FUNCTION "LGF_IntToString" : String   // FC10046, SCL
{ S7_Optimized_Access := 'TRUE' }
VERSION : 0.1
   VAR_INPUT
      intValue : DInt;   // Integer value to convert
   END_VAR
   VAR_TEMP
      tempString : String;   // Temp string
   END_VAR
   // Ret_Val : Converted integer
BEGIN
   //=============================================================================
   // Siemens AG
   // (c)Copyright 2017
   //-----------------------------------------------------------------------------
   // Library:       LGF (Library General Functions)
   // Tested with:   CPU1212C DC/DC/DC FW:V4.2
   // Engineering:   TIA Portal V14 SP1 Upd 5
   // Restrictions:  -
   // Requirements:  PLC (S7-1200 / S7-1500)
   // Functionality: This function converts a integer value to a string
   //-----------------------------------------------------------------------------
   // Change log table:
   // Version  Date        In charge / Changes applied
   // 01.00.00 04.07.2018  Siemens Industry Online Support
   //                      First released version
   // 01.00.01 17.08.2018  Siemens Industry Online Support
   //                      Upgrade: TIA V15 Update 2
   // 01.00.02 23.11.2018  Siemens Industry Online Support
   //                      Upgrade: TIA V15.1
   //=============================================================================

   // Convert integer to string
   #tempString := DINT_TO_STRING(#intValue);

   // Delete padding before number
   WHILE (FIND(IN1 := #tempString, IN2 := ' ') <> 0) DO
     #tempString := DELETE(IN := #tempString, L := 1, P := 1);
   END_WHILE;

   // Output string
   #LGF_IntToString := #tempString;
END_FUNCTION

FUNCTION "LGF_UnixTimeToDTL" : DTL   // FC10047, SCL
{ S7_Optimized_Access := 'TRUE' }
VERSION : 0.1
   VAR_INPUT
      timeUnix : DInt;   // Unix time to convert
   END_VAR
   VAR_OUTPUT
      error : Bool;   // Error = TRUE: Time is outside of allowed range
   END_VAR
   VAR_TEMP
      tempDate : DInt;   // Temporary Date value
      tempTime : DInt;   // Temporary Time value
      tempDTL : DTL;   // Temporary DTL value
   END_VAR
   // Ret_Val : Converted time in DTL
   VAR CONSTANT
      DELTA_1970_1990 : DInt := 631_152_000;   // Delta between 1970-1-1 and 1990-1-1 in seconds (IEC Time Base)
      SEC_PER_DAY : DInt := 86400;   // 86400 seconds in 1 day
   END_VAR
BEGIN
   //=============================================================================
   // Siemens AG
   // (c)Copyright 2017
   //-----------------------------------------------------------------------------
   // Library:       LGF (Library General Functions)
   // Tested with:   CPU1212C DC/DC/DC FW:V4.2
   // Engineering:   TIA Portal V15
   // Restrictions:  -
   // Requirements:  PLC (S7-1200 / S7-1500)
   // Functionality: This function converts Unix time to DTL
   //-----------------------------------------------------------------------------
   // Change log table:
   // Version  Date        In charge / Changes applied
   // 01.00.00 16.10.2018  Siemens Industry Online Support
   //                      First released version
   //=============================================================================

   #error := FALSE;

   // Check if timeUnix less than 01.01.1990
   IF (#timeUnix < #DELTA_1970_1990)
   THEN
     #error := TRUE;
     #LGF_UnixTimeToDTL := DTL#1990-01-01-00:00:00;
     RETURN;
   END_IF;

   // Convert date
   #tempDate := (#timeUnix - #DELTA_1970_1990) / #SEC_PER_DAY;
   #tempDTL := DATE_TO_DTL(DINT_TO_DATE(#tempDate));

   // Convert time
   #tempTime := #timeUnix - #DELTA_1970_1990 - (#tempDate * #SEC_PER_DAY);
   #tempDTL.HOUR := DINT_TO_USINT(#tempTime / 3600);
   #tempDTL.MINUTE := DINT_TO_USINT(#tempTime MOD 3600 / 60);
   #tempDTL.SECOND := DINT_TO_USINT(#tempTime MOD 60);

   // Output date and time
   #LGF_UnixTimeToDTL := #tempDTL;
END_FUNCTION

FUNCTION "LGF_DTLToUnixTime" : DInt   // FC10048, SCL
{ S7_Optimized_Access := 'TRUE' }
VERSION : 0.1
   VAR_INPUT
      timeDTL : DTL;   // Time in DTL to convert
   END_VAR
   VAR_OUTPUT
      error : Bool;   // Error = TRUE: Time is outside of allowed range
   END_VAR
   // Ret_Val : Converted Unix time
   VAR CONSTANT
      DELTA_1970_1990 : DInt := 631_152_000;   // Delta between 1970-1-1 and 1990-1-1 in seconds (IEC Time Base)
      SEC_PER_DAY : DInt := 86400;   // 86400 seconds in 1 day
   END_VAR
BEGIN
   //=============================================================================
   // Siemens AG
   // (c)Copyright 2017
   //-----------------------------------------------------------------------------
   // Library:       LGF (Library General Functions)
   // Tested with:   CPU1212C DC/DC/DC FW:V4.2
   // Engineering:   TIA Portal V15
   // Restrictions:  -
   // Requirements:  PLC (S7-1200 / S7-1500)
   // Functionality: This function converts DTL to Unix time
   //-----------------------------------------------------------------------------
   // Change log table:
   // Version  Date        In charge / Changes applied
   // 01.00.00 16.10.2018  Siemens Industry Online Support
   //                      First released version
   //=============================================================================

   #error := FALSE;

   // Check if timeUnix less than 01.01.1990
   IF (#timeDTL < DTL#1990-01-01-00:00:00)
   THEN
     #error := TRUE;
     #LGF_DTLToUnixTime := 0;
     RETURN;
   END_IF;

   // Convert System Time (UTC) to UNIX time
   #LGF_DTLToUnixTime := (DATE_TO_DINT(DTL_TO_DATE(#timeDTL)) * #SEC_PER_DAY)
                       + (TOD_TO_DINT(DTL_TO_TOD(#timeDTL)) / 1000)
                       + #DELTA_1970_1990;
END_FUNCTION

// folder: Phisical_functions/LGF/7 Signal generators

FUNCTION_BLOCK "LGF_Frequency"   // FB10024, SCL
{ S7_Optimized_Access := 'TRUE' }
   VAR_INPUT
      frequency : Real;   // Input in Hz
      pulsePauseRatio : Real := 1.0;   // Pulse pause ratio
   END_VAR
   VAR_OUTPUT
      clock : Bool;   // -
      countdown : Time;   // -
   END_VAR
   VAR
      instTofTimePulse : TOF_TIME;   // -
      instTofTimePause : TOF_TIME;   // -
      statFrequency : Real;   // -
      statTimePeriod : Time;   // -
      statTimePulse : Time;   // -
      statTimePause : Time;   // -
      statPulsePauseRatio : Real;   // -
   END_VAR
   VAR_TEMP
      tempPulseRate : Real;   // -
      tempPauseRate : Real;   // -
   END_VAR
   VAR CONSTANT
      NULL : Real := 0.0;   // -
   END_VAR
BEGIN
   //=============================================================================
   // SIEMENS AG
   // (c)Copyright 2017
   //-----------------------------------------------------------------------------
   // Library:       LGF (Library General Functions)
   // Tested with:   CPU1214C DC/DC/DC FW:V4.2
   // Engineering:   TIA Portal V14
   // Restrictions:  -
   // Requirements:  PLC (S7-1200, S7-1500)
   // Functionality: Generates frequency signal
   //-----------------------------------------------------------------------------
   // Change log table:
   // Version  Date        Expert in charge / Changes applied
   // 01.00.00 19.08.2015  Siemens Industry Online Support
   //                      First released version
   // 01.01.00 25.05.2016  Siemens Industry Online Support
   //                      New function: pulse pause ratio
   // 01.01.01 26.05.2016  Siemens Industry Online Support
   //                      Add comments
   // 01.01.02 02.01.2017  Siemens Industry Online Support
   //                      Upgrade: TIA Portal V14 Update 1
   // 01.01.03 17.08.2018  Siemens Industry Online Support
   //                      Upgrade: TIA V15 Update 2
   // 01.01.04 23.11.2018  Siemens Industry Online Support
   //                      Upgrade: TIA V15.1
   //=============================================================================

   IF (#frequency <= #NULL) OR (#pulsePauseRatio <= #NULL)  // If input is <= 0.0 : block is off
   THEN
     #clock := FALSE;
     #countdown := t#0s;
   ELSE
     // assign frequency and pulse pause ratio one time 
     IF #statFrequency <> #frequency OR #statPulsePauseRatio <> #pulsePauseRatio THEN
       RESET_TIMER(TIMER := #instTofTimePause);
       RESET_TIMER(TIMER := #instTofTimePulse);

       #tempPulseRate := #pulsePauseRatio / (#pulsePauseRatio + 1); // Calculate pulse rate   
       #tempPauseRate := 1.0 - #tempPulseRate;                      // Calculate pause rate   
       #statTimePeriod := UDINT_TO_TIME(REAL_TO_UDINT((1000.0 / #frequency)));                 // Calculate period time 
       #statTimePulse := UDINT_TO_TIME(REAL_TO_UDINT((1000.0 * #tempPulseRate / #frequency))); // Calculate pulse time   
       #statTimePause := UDINT_TO_TIME(REAL_TO_UDINT((1000.0 * #tempPauseRate / #frequency))); // Calculate pause time
       #statFrequency := #frequency;
       #statPulsePauseRatio := #pulsePauseRatio;
     END_IF;

     // TOF_off expired >> Start again
     #instTofTimePulse(IN := NOT #instTofTimePause.Q,
                       PT := #statTimePulse);
     #countdown := #statTimePulse - #instTofTimePulse.ET;

     #instTofTimePause(IN := #instTofTimePulse.Q,
                       PT := #statTimePause);

     IF #countdown = t#0s THEN
       #countdown := #statTimePause - #instTofTimePause.ET;
     END_IF;

     #clock := #instTofTimePulse.Q; // Assign ouptut 
   END_IF;
END_FUNCTION_BLOCK

FUNCTION_BLOCK "LGF_Impulse"   // FB10025, SCL
{ S7_Optimized_Access := 'TRUE' }
   VAR_INPUT
      frequency : Real;   // Frequnency in Hz
   END_VAR
   VAR_OUTPUT
      impulse : Bool;   // Impulse output
      countdown : Time;   // -
   END_VAR
   VAR
      instTofTimePulse : TOF_TIME;
      statFrequency : Real;
      statTimePulse : Time;
   END_VAR
   VAR_TEMP
      tempImpulse : Bool;
      tempCountdown : Time;
   END_VAR
BEGIN
   //=============================================================================
   // SIEMENS AG
   // (c)Copyright 2017
   //-----------------------------------------------------------------------------
   // Library:       LGF (Library General Functions)
   // Tested with:   CPU1212C DC/DC/DC FW:V4.1
   // Engineering:   TIA Portal V14 Update 1
   // Restrictions:  -
   // Requirements:  PLC (S7-1200 / S7-1500)
   // Functionality: This fuction block generates impulses in the given frequency 
   //-----------------------------------------------------------------------------
   // Change log table:
   // Version  Date        Expert in charge / Changes applied
   // 01.00.00 19.08.2015  Siemens Industry Online Support
   //                      First released version
   // 01.01.01 16.06.2015  Siemens Industry Online Support
   //                      LGF_Impulse calls new LGF_Frequency V1.1.1
   // 01.01.02 02.01.2017  Siemens Industry Online Support
   //                      Upgrade: TIA Portal V14 Update 1
   // 01.02.00 02.02.2017  Siemens Industry Online Support
   //                      Code optimization: no call of LGF_Frequency
   //                      Fix at output "countdown"
   // 01.02.01 17.08.2018  Siemens Industry Online Support
   //                      Upgrade: TIA V15 Update 2
   // 01.02.02 23.11.2018  Siemens Industry Online Support
   //                      Upgrade: TIA V15.1
   //=============================================================================

   IF #frequency <= 0.0 THEN
     #tempImpulse := FALSE;
     #tempCountdown := t#0s;

   ELSE
     // Assign frequency
     #statTimePulse := t#1000s / TRUNC(#frequency * 1000);
     #statFrequency := #frequency;

     // Assign impulse
     #tempImpulse := NOT #instTofTimePulse.Q;

     // Time pulse expired >> Start again
     #instTofTimePulse(IN := NOT #instTofTimePulse.Q,
                       PT := #statTimePulse);

     // Assign countdown
     #tempCountdown := #statTimePulse - #instTofTimePulse.ET;
   END_IF;

   // Write outputs
   #impulse := #tempImpulse;
   #countdown := #tempCountdown;
END_FUNCTION_BLOCK

FUNCTION_BLOCK "LGF_SawTooth"   // FB10026, SCL
{ S7_Optimized_Access := 'TRUE' }
   VAR_INPUT
      startValue : Int;
      timeRange : Time;
      incrementRange : Int;
      numberSteps : Int;
      endlessSteps : Bool;
      restart : Bool;
   END_VAR
   VAR_OUTPUT
      value : Int;
   END_VAR
   VAR
      statStartValue : Int;   // start value of the saw tooth
      statTimeRange : Time;   // time of one period
      statIncrementRange : Int;   // difference from one to another value
      statNumberSteps : Int;   // number of steps
      statEndlessSteps : Bool;
      statCurrentStep : Int;
      statPrevValue : Int;
      statFirstRun : Bool := TRUE;
      statEndlessOn : Bool;
      statStartTimer : Bool;
      statTimerFinished : Bool;
      instTimer : TON_TIME;
      statActValue : Int;
   END_VAR
BEGIN
   //=============================================================================
   // SIEMENS AG
   // (c)Copyright 2017
   //-----------------------------------------------------------------------------
   // Library:       LGF(Library General Functions)
   // Tested with:   CPU1212C DC/DC/DC FW:V4.2
   // Engineering:   TIA Portal V14 Update 1
   // Restrictions:  -
   // Requirements:  PLC (S7-1200 / S7-1500)
   // Functionality: Saw tooth generator
   //-----------------------------------------------------------------------------
   // Change log table:
   // Version  Date        Expert in charge / Changes applied
   // 01.00.00 19.08.2015  Siemens Industry Online Support
   //                      First released version
   // 01.00.01 02.11.2015  Siemens Industry Online Support
   //                      Bug fix
   // 01.00.02 02.01.2017  Siemens Industry Online Support
   //                      Upgrade: TIA Portal V14 Update 1
   // 01.00.03 17.08.2018  Siemens Industry Online Support
   //                      Upgrade: TIA V15 Update 2
   // 01.00.04 23.11.2018  Siemens Industry Online Support
   //                      Upgrade: TIA V15.1
   //=============================================================================

   // Initialization for the first call or reset complete function
   IF (#statFirstRun = TRUE)
     OR (#restart = TRUE) THEN

     // Copy all input parameter to static values
     #statStartValue := #startValue;
     #statTimeRange := #timeRange;
     #statIncrementRange := #incrementRange;
     #statNumberSteps := #numberSteps;
     #statEndlessSteps := #endlessSteps;

     // Reset static values
     #statActValue := #statStartValue;
     #statStartTimer := TRUE;
     #statCurrentStep := 0;
     #statFirstRun := FALSE;
   END_IF;

   // Calculation of a new values if the time base is up
   IF #statTimerFinished = TRUE
     AND (#restart = FALSE) THEN

     #statActValue := #statActValue + #statIncrementRange;
     #statCurrentStep := #statCurrentStep + 1;

     // If a defined number of steps must be performed 
     IF (#statEndlessSteps = FALSE) THEN

       // Restart with start value if number of steps is reached
       IF #statCurrentStep > #statNumberSteps THEN

         #statCurrentStep := 0;
         #statActValue := #statStartValue;
       END_IF;

       // If endless is on the step counter is resetted  
     ELSE

       #statEndlessOn := TRUE;
       #statCurrentStep := 0;
     END_IF;

     #statStartTimer := FALSE; // Reset the time base
   END_IF;

   // Call a times as basis of the step range
   #instTimer(IN := #statStartTimer,
              PT := #statTimeRange,
              Q => #statTimerFinished);

   // Start the timer
   #statStartTimer := TRUE;

   // Write Output, if restart is active output value = 0
   IF (#restart = TRUE) THEN
     #statActValue := #startValue;
   END_IF;

   #value := #statActValue;
END_FUNCTION_BLOCK

FUNCTION_BLOCK "LGF_SinusCI"   // FB10027, SCL
{ S7_Optimized_Access := 'TRUE' }
VERSION : 0.1
   VAR_INPUT
      amplitude : Real := 0.0;   // Amplitude
      offset : Real := 1000.0;   // Offset
      periodeMS : UDInt := 1000;   // Periode in milliseconds
      callOB : OB_Cyclic;   // Call OB
      reset : Bool;   // Reset values
   END_VAR
   VAR_OUTPUT
      sinusValues : Real;   // Calculated Sinus values
      error : Bool;   // "0" = no error; "1" = error
      statusID : UInt;   // Error source
      status : Word;   // Status and error codes
   END_VAR
   VAR
      statRad : Real;   // Size of an angle in radians
      statCounter : UDInt;   // Counter value
   END_VAR
   VAR_TEMP
      tempCycleTime : UDInt;   // Temp cycle time from CallOB
      tempCyclePhase : UDInt;   // Temp cycle phase from CallOB
      tempCycleStatus : Word;   // Temp cycle status from CallOB
      tempReadTimeStatus : Int;   // Return value of QRY_CINT
   END_VAR
   VAR CONSTANT
      PI : Real := 3.141593;   // PI
      NO_ERROR : Word := 16#0000;   // Status no error
      OB_UNAVAILABLE : Word := 16#8200;   // Status OB not available
      ERROR_IN_THIS_BLOCK : UInt := 1;   // Error ID local error
      ERROR_QRY_CINT : UInt := 2;   // Error ID error in function QRY_CINT
   END_VAR
BEGIN
   //=============================================================================
   // Siemens AG
   // (c)Copyright 2017
   //-----------------------------------------------------------------------------
   // Library:       LGF (Library General Functions)
   // Tested with:   CPU1212C DC/DC/DC FW:V4.2
   // Engineering:   TIA Portal V15 Upd 2
   // Restrictions:  -
   // Requirements:  PLC (S7-1200 / S7-1500)
   // Functionality: This function generates a sinus signal
   //-----------------------------------------------------------------------------
   // Change log table:
   // Version  Date        In charge/Changes applied
   // 01.00.00 03.07.2018  Siemens Industry Online Support
   //                      First released version
   // 01.00.01 17.08.2018  Siemens Industry Online Support
   //                      Upgrade: TIA V15 Update 2
   // 01.00.02 23.11.2018  Siemens Industry Online Support
   //                      Upgrade: TIA V15.1
   //-----------------------------------------------------------------------------
   //Status Codes: -
   //=============================================================================

   // Initialize
   #error := FALSE;
   #statusID := #ERROR_IN_THIS_BLOCK;
   #status := #NO_ERROR;

   // get sample time, according to the cyclic interrupt OB number
   #tempReadTimeStatus := QRY_CINT(OB_NR := #callOB, CYCLE => #tempCycleTime,
                                   PHASE => #tempCyclePhase, STATUS => #tempCycleStatus);

   // Generate error message of the QRY_CINT function
   IF (#tempReadTimeStatus <> 0)
   THEN
     #error := TRUE;
     #statusID := #ERROR_QRY_CINT;
     #status := INT_TO_WORD(#tempReadTimeStatus);
     RETURN;
   END_IF;

   // Generate error message when OB unavailable
   IF (#tempCycleStatus = 16#0000)
   THEN
     #error := TRUE;
     #statusID := #ERROR_IN_THIS_BLOCK;
     #status := #OB_UNAVAILABLE;
     RETURN;
   END_IF;

   IF (#reset = TRUE)
   THEN
     #statCounter := 0;
     #sinusValues := 0;
   ELSE
     // Increment Counter with each call of "OB_Cyclic_interrupt"
     #statCounter := #statCounter + (#tempCycleTime) / 1000;
     #statCounter := #statCounter MOD (#periodeMS);

     #statRad := UDINT_TO_REAL(#statCounter) * 2.0 * #PI / (UDINT_TO_REAL(#periodeMS));

     #sinusValues := SIN(#statRad) * #amplitude + #offset;
   END_IF;
END_FUNCTION_BLOCK

FUNCTION_BLOCK "LGF_CosinusCI"   // FB10028, SCL
{ S7_Optimized_Access := 'TRUE' }
VERSION : 0.1
   VAR_INPUT
      amplitude : Real := 0.0;   // Amplitude
      offset : Real := 1000.0;   // Offset
      periodeMS : UDInt := 1000;   // Periode in milliseconds
      callOB : OB_Cyclic;   // Call OB
      reset : Bool;   // Reset values
   END_VAR
   VAR_OUTPUT
      cosinusValues : Real;   // Calculated Cosinus values
      error : Bool;   // "0" = no error; "1" = error
      statusID : UInt;   // Error source
      status : Word;   // Status and error codes
   END_VAR
   VAR
      statRad : Real;   // Size of an angle in radians
      statCounter : UDInt;   // Counter value
   END_VAR
   VAR_TEMP
      tempCycleTime : UDInt;   // Temp cycle time from CallOB
      tempCyclePhase : UDInt;   // Temp cycle phase from CallOB
      tempCycleStatus : Word;   // Temp cycle status from CallOB
      tempReadTimeStatus : Int;   // Return value of QRY_CINT
   END_VAR
   VAR CONSTANT
      PI : Real := 3.141593;   // PI
      NO_ERROR : Word := 16#0000;   // Status no error
      OB_UNAVAILABLE : Word := 16#8200;   // Status OB not available
      ERROR_IN_THIS_BLOCK : UInt := 1;   // Error ID local error
      ERROR_QRY_CINT : UInt := 2;   // Error ID error in function QRY_CINT
   END_VAR
BEGIN
   //=============================================================================
   // Siemens AG
   // (c)Copyright 2017
   //-----------------------------------------------------------------------------
   // Library:       LGF (Library General Functions)
   // Tested with:   CPU1212C DC/DC/DC FW:V4.2
   // Engineering:   TIA Portal V15 Upd 2
   // Restrictions:  -
   // Requirements:  PLC (S7-1200 / S7-1500)
   // Functionality: This function generates a cosinus signal
   //-----------------------------------------------------------------------------
   // Change log table:
   // Version  Date        In charge/Changes applied
   // 01.00.00 03.07.2018  Siemens Industry Online Support
   //                      First released version
   // 01.00.01 17.08.2018  Siemens Industry Online Support
   //                      Upgrade: TIA V15 Update 2
   // 01.00.02 23.11.2018  Siemens Industry Online Support
   //                      Upgrade: TIA V15.1
   //-----------------------------------------------------------------------------
   //Status Codes: -
   //=============================================================================

   // Initialize
   #error := FALSE;
   #statusID := #ERROR_IN_THIS_BLOCK;
   #status := #NO_ERROR;

   // get sample time, according to the cyclic interrupt OB number
   #tempReadTimeStatus := QRY_CINT(OB_NR := #callOB, CYCLE => #tempCycleTime,
                                   PHASE => #tempCyclePhase, STATUS => #tempCycleStatus);

   // Generate error message of the QRY_CINT function
   IF (#tempReadTimeStatus <> 0)
   THEN
     #error := TRUE;
     #statusID := #ERROR_QRY_CINT;
     #status := INT_TO_WORD(#tempReadTimeStatus);
     RETURN;
   END_IF;

   // Generate error message when OB unavailable
   IF (#tempCycleStatus = 16#0000)
   THEN
     #error := TRUE;
     #statusID := #ERROR_IN_THIS_BLOCK;
     #status := #OB_UNAVAILABLE;
     RETURN;
   END_IF;

   IF (#reset = TRUE) 
   THEN
     #statCounter := 0;
     #cosinusValues := 0;
   ELSE
     // Increment Counter with each call of "OB_Cyclic_interrupt"
     #statCounter := #statCounter + (#tempCycleTime) / 1000;
     #statCounter := #statCounter MOD (#periodeMS);

     #statRad := UDINT_TO_REAL(#statCounter) * 2.0 * #PI / (UDINT_TO_REAL(#periodeMS));

     #cosinusValues := COS(#statRad) * #amplitude + #offset;
   END_IF;
END_FUNCTION_BLOCK

FUNCTION_BLOCK "LGF_RectangleCI"   // FB10029, SCL
{ S7_Optimized_Access := 'TRUE' }
VERSION : 0.1
   VAR_INPUT
      amplitude : Real := 0.0;   // Amplitude
      offset : Real := 1000.0;   // Offset
      periodeMS : UDInt := 1000;   // Periode in milliseconds
      callOB : OB_Cyclic;   // Call OB
      reset : Bool;   // Reset values
   END_VAR
   VAR_OUTPUT
      rectangleValues : Real;   // Calculated rectangle values
      error : Bool;   // "0" = no error; "1" = error
      statusID : UInt;   // Error source
      status : Word;   // Status and error codes
   END_VAR
   VAR
      statRad : Real;   // Size of an angle in radians
      statCounter : UDInt;   // Counter value
   END_VAR
   VAR_TEMP
      tempCycleTime : UDInt;   // Temp cycle time from CallOB
      tempCyclePhase : UDInt;   // Temp cycle phase from CallOB
      tempCycleStatus : Word;   // Temp cycle status from CallOB
      tempReadTimeStatus : Int;   // Return value of QRY_CINT
   END_VAR
   VAR CONSTANT
      PI : Real := 3.141593;   // PI
      NO_ERROR : Word := 16#0000;   // Status no error
      OB_UNAVAILABLE : Word := 16#8200;   // Status OB not available
      ERROR_IN_THIS_BLOCK : UInt := 1;   // Error ID local error
      ERROR_QRY_CINT : UInt := 2;   // Error ID error in function QRY_CINT
   END_VAR
BEGIN
   //=============================================================================
   // Siemens AG
   // (c)Copyright 2017
   //-----------------------------------------------------------------------------
   // Library:       LGF (Library General Functions)
   // Tested with:   CPU1212C DC/DC/DC FW:V4.2
   // Engineering:   TIA Portal V15 Upd 2
   // Restrictions:  -
   // Requirements:  PLC (S7-1200 / S7-1500)
   // Functionality: This function generates a rectangle signal
   //-----------------------------------------------------------------------------
   // Change log table:
   // Version  Date        In charge/Changes applied
   // 01.00.00 03.07.2018  Siemens Industry Online Support
   //                      First released version
   // 01.00.01 17.08.2018  Siemens Industry Online Support
   //                      Upgrade: TIA V15 Update 2
   // 01.00.02 23.11.2018  Siemens Industry Online Support
   //                      Upgrade: TIA V15.1
   //-----------------------------------------------------------------------------
   //Status Codes: -
   //=============================================================================

   // Initialize
   #error := FALSE;
   #statusID := #ERROR_IN_THIS_BLOCK;
   #status := #NO_ERROR;

   // get sample time, according to the cyclic interrupt OB number
   #tempReadTimeStatus := QRY_CINT(OB_NR := #callOB, CYCLE => #tempCycleTime,
                                   PHASE => #tempCyclePhase, STATUS => #tempCycleStatus);

   // Generate error message of the QRY_CINT function
   IF (#tempReadTimeStatus <> 0)
   THEN
     #error := TRUE;
     #statusID := #ERROR_QRY_CINT;
     #status := INT_TO_WORD(#tempReadTimeStatus);
     RETURN;
   END_IF;

   // Generate error message when OB unavailable
   IF (#tempCycleStatus = 16#0000)
   THEN
     #error := TRUE;
     #statusID := #ERROR_IN_THIS_BLOCK;
     #status := #OB_UNAVAILABLE;
     RETURN;
   END_IF;

   IF (#reset = TRUE) 
   THEN
     #statCounter := 0;
     #rectangleValues := 0;
   ELSE
     // Increment Counter with each call of "OB_Cyclic_interrupt"
     #statCounter := #statCounter + (#tempCycleTime) / 1000;
     #statCounter := #statCounter MOD (#periodeMS);

     IF (#statCounter <= (#periodeMS / 2))
     THEN
       #rectangleValues := #offset + #amplitude;
     ELSE
       #rectangleValues := #offset - #amplitude;
     END_IF;
   END_IF;
END_FUNCTION_BLOCK

FUNCTION_BLOCK "LGF_TriangleCI"   // FB10030, SCL
{ S7_Optimized_Access := 'TRUE' }
VERSION : 0.1
   VAR_INPUT
      amplitude : Real := 0.0;   // Amplitude
      offset : Real := 1000.0;   // Offset
      periodeMS : UDInt := 1000;   // Periode in milliseconds
      callOB : OB_Cyclic;   // Call OB
      reset : Bool;   // Reset values
   END_VAR
   VAR_OUTPUT
      triangleValues : Real;   // Calculated triangle values
      error : Bool;   // "0" = no error; "1" = error
      statusID : UInt;   // Error source
      status : Word;   // Status and error codes
   END_VAR
   VAR
      statRad : Real;   // Size of an angle in radians
      statCounter : UDInt;   // Counter value
   END_VAR
   VAR_TEMP
      tempCycleTime : UDInt;   // Temp cycle time from CallOB
      tempCyclePhase : UDInt;   // Temp cycle phase from CallOB
      tempCycleStatus : Word;   // Temp cycle status from CallOB
      tempReadTimeStatus : Int;   // Return value of QRY_CINT
   END_VAR
   VAR CONSTANT
      PI : Real := 3.141593;   // PI
      NO_ERROR : Word := 16#0000;   // Status no error
      OB_UNAVAILABLE : Word := 16#8200;   // Status OB not available
      ERROR_IN_THIS_BLOCK : UInt := 1;   // Error ID local error
      ERROR_QRY_CINT : UInt := 2;   // Error ID error in function QRY_CINT
   END_VAR
BEGIN
   //=============================================================================
   // Siemens AG
   // (c)Copyright 2017
   //-----------------------------------------------------------------------------
   // Library:       LGF (Library General Functions)
   // Tested with:   CPU1212C DC/DC/DC FW:V4.2
   // Engineering:   TIA Portal V15 Upd 2
   // Restrictions:  -
   // Requirements:  PLC (S7-1200 / S7-1500)
   // Functionality: This function generates a rectangle signal
   //-----------------------------------------------------------------------------
   // Change log table:
   // Version  Date        In charge/Changes applied
   // 01.00.00 03.07.2018  Siemens Industry Online Support
   //                      First released version
   // 01.00.01 17.08.2018  Siemens Industry Online Support
   //                      Upgrade: TIA V15 Update 2
   // 01.00.02 23.11.2018  Siemens Industry Online Support
   //                      Upgrade: TIA V15.1
   //-----------------------------------------------------------------------------
   //Status Codes: -
   //=============================================================================

   // Initialize
   #error := FALSE;
   #statusID := #ERROR_IN_THIS_BLOCK;
   #status := #NO_ERROR;

   // get sample time, according to the cyclic interrupt OB number
   #tempReadTimeStatus := QRY_CINT(OB_NR := #callOB, CYCLE => #tempCycleTime,
                                   PHASE => #tempCyclePhase, STATUS => #tempCycleStatus);

   // Generate error message of the QRY_CINT function
   IF (#tempReadTimeStatus <> 0)
   THEN
     #error := TRUE;
     #statusID := #ERROR_QRY_CINT;
     #status := INT_TO_WORD(#tempReadTimeStatus);
     RETURN;
   END_IF;

   // Generate error message when OB unavailable
   IF #tempCycleStatus = 16#0000 THEN
     #error := TRUE;
     #statusID := #ERROR_IN_THIS_BLOCK;
     #status := #OB_UNAVAILABLE;
     RETURN;
   END_IF;

   IF (#reset = TRUE) 
   THEN
     #statCounter := 0;
     #triangleValues := 0;
   ELSE
     // Increment Counter with each call of "OB_Cyclic_interrupt"
     #statCounter := #statCounter + (#tempCycleTime) / 1000;
     #statCounter := #statCounter MOD (#periodeMS);

     IF (#statCounter <= (#periodeMS / 2))
     THEN
       #triangleValues := 4.0 * #amplitude /  UDINT_TO_REAL(#periodeMS) * UDINT_TO_REAL(#statCounter)  - #amplitude + #offset;
     ELSE
       #triangleValues := -4.0 * #amplitude / UDINT_TO_REAL(#periodeMS) * UDINT_TO_REAL(#statCounter) + 3 * #amplitude + #offset;
     END_IF;
   END_IF;
END_FUNCTION_BLOCK

FUNCTION_BLOCK "LGF_SawToothCI"   // FB10031, SCL
{ S7_Optimized_Access := 'TRUE' }
VERSION : 0.1
   VAR_INPUT
      amplitude : Real := 0.0;   // Amplitude
      offset : Real := 1000.0;   // Offset
      periodeMS : UDInt := 1000;   // Periode in milliseconds
      callOB : OB_Cyclic;   // Call OB
      reset : Bool;   // Reset values
   END_VAR
   VAR_OUTPUT
      sawToothValues : Real;   // Calculated saw tooth values
      error : Bool;   // "0" = no error; "1" = error
      statusID : UInt;   // Error source
      status : Word;   // Status and error codes
   END_VAR
   VAR
      statRad : Real;   // Size of an angle in radians
      statCounter : UDInt;   // Counter value
   END_VAR
   VAR_TEMP
      tempCycleTime : UDInt;   // Temp cycle time from CallOB
      tempCyclePhase : UDInt;   // Temp cycle phase from CallOB
      tempCycleStatus : Word;   // Temp cycle status from CallOB
      tempReadTimeStatus : Int;   // Return value of QRY_CINT
   END_VAR
   VAR CONSTANT
      PI : Real := 3.141593;   // PI
      NO_ERROR : Word := 16#0000;   // Status no error
      OB_UNAVAILABLE : Word := 16#8200;   // Status OB not available
      ERROR_IN_THIS_BLOCK : UInt := 1;   // Error ID local error
      ERROR_QRY_CINT : UInt := 2;   // Error ID error in function QRY_CINT
   END_VAR
BEGIN
   //=============================================================================
   // Siemens AG
   // (c)Copyright 2017
   //-----------------------------------------------------------------------------
   // Library:       LGF (Library General Functions)
   // Tested with:   CPU1212C DC/DC/DC FW:V4.2
   // Engineering:   TIA Portal V15 Upd 2
   // Restrictions:  -
   // Requirements:  PLC (S7-1200 / S7-1500)
   // Functionality: This function generates a rectangle signal
   //-----------------------------------------------------------------------------
   // Change log table:
   // Version  Date        In charge/Changes applied
   // 01.00.00 03.07.2018  Siemens Industry Online Support
   //                      First released version
   // 01.00.01 17.08.2018  Siemens Industry Online Support
   //                      Upgrade: TIA V15 Update 2
   // 01.00.02 23.11.2018  Siemens Industry Online Support
   //                      Upgrade: TIA V15.1
   //-----------------------------------------------------------------------------
   //Status Codes: -
   //=============================================================================

   // Initialize
   #error := FALSE;
   #statusID := #ERROR_IN_THIS_BLOCK;
   #status := #NO_ERROR;

   // get sample time, according to the cyclic interrupt OB number
   #tempReadTimeStatus := QRY_CINT(OB_NR := #callOB, CYCLE => #tempCycleTime,
                                   PHASE => #tempCyclePhase, STATUS => #tempCycleStatus);

   // Generate error message of the QRY_CINT function
   IF (#tempReadTimeStatus <> 0)
   THEN
     #error := TRUE;
     #statusID := #ERROR_QRY_CINT;
     #status := INT_TO_WORD(#tempReadTimeStatus);
     RETURN;
   END_IF;

   // Generate error message when OB unavailable
   IF (#tempCycleStatus = 16#0000)
   THEN
     #error := TRUE;
     #statusID := #ERROR_IN_THIS_BLOCK;
     #status := #OB_UNAVAILABLE;
     RETURN;
   END_IF;

   IF (#reset = TRUE)
   THEN
     #statCounter := 0;
     #sawToothValues := 0;
   ELSE
     // Increment Counter with each call of "OB_Cyclic_interrupt"
     #statCounter := #statCounter + (#tempCycleTime) / 1000;
     #statCounter := #statCounter MOD (#periodeMS);

     #sawToothValues := 2.0 * #amplitude / UDINT_TO_REAL(#periodeMS) * UDINT_TO_REAL(#statCounter) - #amplitude + #offset;

   END_IF;
END_FUNCTION_BLOCK

// folder: Phisical_functions/LGF/8 Technology operations

FUNCTION_BLOCK "LGF_LimRateOfChangeBasic"   // FB10032, SCL
{ S7_Optimized_Access := 'TRUE' }
VERSION : 0.1
   VAR_INPUT
      inputValue : Real;   // Input Value/ setpoint
      setRateLim : Real;   // rate of change limitation (1/second)
      defaultOutValue : Real;   // default output value
      onDefaultOutValue : Bool;   // default output value on (outputValue=defaultOutValue)
      callOB : OB_Cyclic;   // cyclic interrupt OB
   END_VAR
   VAR_OUTPUT
      outputValue : Real;   // output value
      error : Bool;   // "0" = no error; "1" = error
      statusID : UInt;   // Error destination: "1" = LGFLimRateOfChangeBasic; "2" = QRY_CINT
      status : Word;   // status and error codes
   END_VAR
   VAR
      statPrevTime : DTL;   // -
      statPrevOut : Real;   // -
   END_VAR
   VAR_TEMP
      tempCycleTime : UDInt;   // -
      tempCylcePhase : UDInt;   // -
      tempCycleStatus : Word;   // -
      tempDeltaTime : Time;   // -
      tempCycleTimeReal : Real;   // -
      tempReadTimeStatus : Int;   // -
      tempOut : Real;   // -
   END_VAR
   VAR CONSTANT
      NO_ERROR : Word := 16#0000;   // -
      INIT_VALUE : Word := 16#7000;   // -
      OB_UNAVAILABLE : Word := 16#8200;   // -
      NEG_RATE_LIM : Word := 16#8201;   // -
      ERROR_IN_THIS_BLOCK : UInt := 1;   // -
      ERROR_QRY_CINT : UInt := 2;   // -
   END_VAR
BEGIN
   //=============================================================================
   // Siemens AG
   // (c)Copyright 2017
   //-----------------------------------------------------------------------------
   // Library:       LGF(Library General Functions)
   // Tested with:   CPU1212C DC/DC/DC FW:V4.2
   // Engineering:   TIA Portal V14 Update 1
   // Restrictions:  only callable in a cyclic interrupt OB
   // Requirements:  PLC (S7-1200 / S7-1500)
   // Functionality: This function block generates a ramp function from a step function.
   //-----------------------------------------------------------------------------
   // Change log table:
   // Version  Date        In charge / Changes applied
   // 01.00.00 21.06.2016  Siemens Industry Online Support
   //                      First released version
   // 01.00.01 02.01.2017  Siemens Industry Online Support
   //                      Upgrade: TIA Portal V14 Update 1
   // 01.00.02 17.08.2018  Siemens Industry Online Support
   //                      Upgrade: TIA V15 Update 2
   // 01.00.03 23.11.2018  Siemens Industry Online Support
   //                      Upgrade: TIA V15.1
   //-----------------------------------------------------------------------------
   //Status Codes:
   // 16#0000:  No errors
   // 16#7000:  Initial value
   // 16#8200:  Call OB unavailable
   // 16#8201:  Negativ value for rate of change
   //=============================================================================

   // Set no errors
   #error := FALSE;
   #statusID := #ERROR_IN_THIS_BLOCK;
   #status := #NO_ERROR;

   // Read cycle time of the call OB
   #tempReadTimeStatus := QRY_CINT(OB_NR := #callOB, CYCLE => #tempCycleTime, PHASE => #tempCylcePhase, STATUS => #tempCycleStatus);
   #tempCycleTimeReal := UDINT_TO_REAL(#tempCycleTime) / 1.0e6;

   // Generate error message of the QRY_CINT function
   IF (#tempReadTimeStatus <> 0) THEN
     #error := TRUE;
     #statusID := #ERROR_QRY_CINT;
     #status := INT_TO_WORD(#tempReadTimeStatus);
     RETURN;
   END_IF;

   // Generate error message when OB unavailable
   IF #tempCycleStatus = 16#0000 THEN
     #error := TRUE;
     #statusID := #ERROR_IN_THIS_BLOCK;
     #status := #OB_UNAVAILABLE;
     RETURN;
   END_IF;

   IF #setRateLim < 0.0 THEN
     #error := TRUE;
     #statusID := #ERROR_IN_THIS_BLOCK;
     #status := #NEG_RATE_LIM;
     RETURN;
   END_IF;

   // Initialize start point
   IF #onDefaultOutValue = true THEN
     #statPrevOut := #defaultOutValue;
     #outputValue := #defaultOutValue;
     #status := #INIT_VALUE;
     RETURN;
   END_IF;

   #tempOut := #statPrevOut;

   // Ramp function
   IF #inputValue < #tempOut THEN
     #tempOut := #tempOut - (#setRateLim * #tempCycleTimeReal);
     #tempOut := MAX(IN1 := #tempOut, IN2 := #inputValue);
     #statPrevOut := #tempOut;
   ELSE
     IF #inputValue > #tempOut THEN
       #tempOut := (#setRateLim * #tempCycleTimeReal) + #tempOut;
       #tempOut := MIN(IN1 := #tempOut, IN2 := #inputValue);
       #statPrevOut := #tempOut;
     END_IF;
   END_IF;

   #outputValue := #tempOut;
END_FUNCTION_BLOCK

FUNCTION_BLOCK "LGF_LimRateOfChangeAdvanced"   // FB10033, SCL
{ S7_Optimized_Access := 'TRUE' }
VERSION : 0.1
   VAR_INPUT
      inputValue : Real;   // input value
      setPosUpRateLim : Real;   // limit up rate of change in positiv range (1/second)
      setPosDownRateLim : Real;   // limit down rate of change in positiv range (1/second)
      setNegUpRateLim : Real;   // limit up rate of change in nagativ range (1/second)
      setNegDownRateLim : Real;   // limit down rate of change in nagativ range (1/second)
      setHighLim : Real;   // high limit
      setLowLim : Real;   // low limit
      processValue : Real;   // process value
      defaultOutValue : Real;   // default output value
      onDefaultOutValue : Bool;   // default output value on (outputValue=defaultOutValue)
      track : Bool;   // tracking (outVal=inputValue)
      manOp : Bool;   // manual mode on (outputValue=processValue)
      reset : Bool;   // complete restart
      callOB : OB_Cyclic;   // cyclic interrupt OB
   END_VAR
   VAR_OUTPUT
      outputValue : Real;   // output value
      posUpRateLim : Bool;   // up rate limit in positiv range reached
      posDownRateLim : Bool;   // down rate limit in positiv range reached
      negUpRateLim : Bool;   // up rate limit in negative range reached
      negDownRateLim : Bool;   // down rate limit in negativ range reached
      highLim : Bool;   // high limit reached
      lowLim : Bool;   // low limit reached
      error : Bool;   // "0" = no error; "1" = error
      statusID : UInt;   // Error destination: "1" = LGFLimRateOfChangeAdvanced; "2" = QRY_CINT
      status : Word;   // status and error codes
   END_VAR
   VAR
      statPrevOutputValue : Real := 0.0;   // -
      statManOp : Bool;   // -
   END_VAR
   VAR_TEMP
      tempPosUp : Bool;   // -
      tempPosDown : Bool;   // -
      tempNegUp : Bool;   // -
      tempNegDown : Bool;   // -
      tempHighLim : Bool;   // -
      tempLowLim : Bool;   // -
      tempCycleReal : Real;   // -
      tempOutv : Real;   // -
      tempVar : Real;   // -
      tempCycleTime : UDInt;   // -
      tempCyclePhase : UDInt;   // -
      tempCycleStatus : Word;   // -
      tempReadTimeStatus : Int;   // -
   END_VAR
   VAR CONSTANT
      NO_ERROR : Word := 16#0000;   // -
      OB_UNAVAILABLE : Word := 16#8200;   // -
      HIGHLIM_UNDER_LOWLIM : Word := 16#8201;   // -
      NEG_RATE_OF_CHANGE : Word := 16#8202;   // -
      ERROR_IN_THIS_BLOCK : UInt := 1;   // -
      ERROR_QRY_CINT : UInt := 2;   // -
   END_VAR
BEGIN
   //=============================================================================
   // Siemens AG
   // (c)Copyright 2017
   //-----------------------------------------------------------------------------
   // Library:       LGF(Library General Functions)
   // Tested with:   CPU1212C DC/DC/DC FW:V4.2
   // Engineering:   TIA Portal V14 Update 1
   // Restrictions:  only callable just in cyclic interrupt OB
   // Requirements:  PLC (S7-1200 / S7-1500)
   // Functionality: This function block generates a ramp function from a step 
   //                function with advanced modes and settings.  
   //-----------------------------------------------------------------------------
   // Change log table:
   // Version  Date        In charge / Changes applied
   // 01.00.00 21.06.2016  Siemens Industry Online Support
   //                      First released version
   // 01.00.01 02.01.2017  Siemens Industry Online Support
   //                      Upgrade: TIA Portal V14 Update 1
   // 01.00.02 17.08.2018  Siemens Industry Online Support
   //                      Upgrade: TIA V15 Update 2
   // 01.00.03 23.11.2018  Siemens Industry Online Support
   //                      Upgrade: TIA V15.1
   //-----------------------------------------------------------------------------
   //Status Codes:
   // 16#0000:  No errors
   // 16#8200:  Call OB unavailable
   // 16#8201:  Paramater for high limit lower thal low limit
   // 16#8202:  Negativ value for the rate of change parameter
   //=============================================================================

   // Initialize
   #error := FALSE;
   #statusID := #ERROR_IN_THIS_BLOCK;
   #status := #NO_ERROR;

   //***// get sample time, according to the cyclic interrupt OB number
   #tempReadTimeStatus := QRY_CINT(OB_NR := #callOB, CYCLE => #tempCycleTime,
                                   PHASE => #tempCyclePhase, STATUS => #tempCycleStatus);
   #tempCycleReal := UDINT_TO_REAL(#tempCycleTime) / 1.0e6; // Time in seconds

   // Generate error message of the QRY_CINT function
   IF (#tempReadTimeStatus <> 0) THEN
     #error := TRUE;
     #statusID := #ERROR_QRY_CINT;
     #status := INT_TO_WORD(#tempReadTimeStatus);
     RETURN;
   END_IF;

   // Generate error message when OB unavailable
   IF #tempCycleStatus = 16#0000 THEN
     #error := TRUE;
     #statusID := #ERROR_IN_THIS_BLOCK;
     #status := #OB_UNAVAILABLE;
     RETURN;
   END_IF;

   IF #setHighLim < #setLowLim THEN
     #error := TRUE;
     #statusID := #ERROR_IN_THIS_BLOCK;
     #status := #HIGHLIM_UNDER_LOWLIM;
     RETURN;
   END_IF;

   IF (#setNegDownRateLim < 0.0) OR (#setNegUpRateLim < 0.0)
     OR (#setPosDownRateLim < 0.0) OR (#setPosUpRateLim < 0.0)
   THEN
     #error := TRUE;
     #statusID := #ERROR_IN_THIS_BLOCK;
     #status := #NEG_RATE_OF_CHANGE;
     RETURN;
   END_IF;

   // Initialize temp variable
   #tempPosUp := FALSE;
   #tempPosDown := FALSE;
   #tempNegUp := FALSE;
   #tempNegDown := FALSE;
   #tempHighLim := FALSE;
   #tempLowLim := FALSE;
   #tempOutv := #inputValue;

   // RESTART
   IF #reset
   THEN
     #statManOp := FALSE;    // reset manual mode flag 
     IF #onDefaultOutValue
       // preset output
     THEN
       #tempOutv := #defaultOutValue;
       // limitation of output
       IF #tempOutv >= #setHighLim
       THEN
         // High limitation
         #tempOutv := #setHighLim;
         #tempHighLim := TRUE;
       END_IF;

       IF #tempOutv <= #setLowLim
       THEN
         // Low limitation
         #tempOutv := #setLowLim;
         #tempLowLim := TRUE;
       END_IF;
     ELSE
       // reset output
       #tempOutv := 0.0;
     END_IF;
   ELSE

     // OPERATING MODES
     // -------------------------------------------------------
     IF #manOp
     THEN
       //---// MANUAL MODE
       // bumples switch between manual mode and auto mode    
       #tempOutv := #processValue;
       // Keep manual mode until setpoint in the space of low and high limit
       #statManOp := TRUE;
     ELSE
       //---// AUTOMATIC MODE
       IF #onDefaultOutValue
       THEN
         // preset output by default value
         #tempOutv := #defaultOutValue;
       ELSE
         IF #track
         THEN
           // output has same value as input
           #tempOutv := #inputValue;
         ELSE
           // REGULAR FUNCTION                    
           // Negativ range
           IF #statPrevOutputValue < 0
           THEN
             IF #statPrevOutputValue > #inputValue
             THEN
               // limited rate of change
               #tempVar := #statPrevOutputValue - #setNegUpRateLim * #tempCycleReal;
               IF #inputValue < #tempVar
               THEN
                 // Setpoint not reached yet
                 // set notification for up rate limit in neg range              
                 #tempNegUp := TRUE;
                 #tempOutv := #tempVar;
               END_IF;
             ELSE
               IF #setNegDownRateLim = 0.0
               THEN
                 // set notification for down rate limit in neg range              
                 #tempNegDown := TRUE;
                 IF #inputValue <= 0.0
                 THEN
                   #tempOutv := #inputValue;
                 ELSE
                   #tempOutv := 0.0;
                 END_IF;
               ELSE
                 IF #inputValue <= 0.0
                 THEN
                   // limited rate of change
                   #tempVar := #statPrevOutputValue + #setNegDownRateLim * #tempCycleReal;
                   IF #inputValue > #tempVar
                   THEN
                     // set notification for down rate limit in neg range
                     #tempNegDown := TRUE;
                     #tempOutv := #tempVar;
                   END_IF;
                 ELSE
                   // changeover between neg. and pos. range
                   // period till zero-crossing
                   #tempVar := - #statPrevOutputValue / #setNegDownRateLim;

                   IF #tempVar <= #tempCycleReal
                   THEN
                     // period till zero-crossing shorten than sample time
                     // limited rate of change
                     #tempVar := (#tempCycleReal - #tempVar) * #setPosUpRateLim;

                     IF #inputValue > #tempVar
                     THEN
                       // set notification for rate limit 
                       #tempNegDown := FALSE;
                       #tempPosUp := TRUE;
                       #tempOutv := #tempVar;
                     END_IF;
                   ELSE
                     // set notification for rate limit
                     #tempNegDown := TRUE;
                     #tempPosUp := FALSE;
                     #tempOutv := #statPrevOutputValue + #tempCycleReal * #setNegDownRateLim;
                   END_IF;
                 END_IF;
               END_IF;
             END_IF;
           ELSE
             // Positiv range + 0                        
             IF #statPrevOutputValue < #inputValue
             THEN
               // limited rate of change
               #tempVar := #statPrevOutputValue + #setPosUpRateLim * #tempCycleReal;
               IF #inputValue > #tempVar
               THEN
                 // set notification for up rate limit in pos range              
                 #tempPosUp := TRUE;
                 #tempOutv := #tempVar;
               END_IF;
             END_IF;